(* Logix 5000 project; controller MV vendor 1 type 14 code 217 rev 31.11; software revision 31.00; part 9 of 53 *)
(* tags used below, declared in another part *)
   MC_CH1_DRAIN : PlantItem;   // CH1_DRAIN
   MC_CH1_LF1 : PlantItem;   // CH1_LF1
   MC_CH1_PR1 : PlantItem;   // CH1_PR1
   MC_CH1_RR : PlantItem;   // CH1_RR
   MC_N100 : INT[255];   // C1_PLC Channel 1 PLC data
   MC_N102 : INT[255];   // CH1 PROG Channel 1 CIP progra m
   MC_N104 : INT[255];   // CH1 REPORT Channel 1 CIP report file
   MC_N112 : INT[255];   // FVR DATA Data read from FV ro uting PLC
   MC_N113 : INT[255];   // MVR DATA Data read from MV ro uting PLC
   MC_N114 : INT[255];   // YP DATA
   MC_N120 : INT[255];   // C2 PLC Channel 2 PLC data
   MC_N80 : INT[255];   // SRV1_PLC Detergent tank 1 ser vice PLC data
   MC_N90 : INT[255];   // SV2_PLC Detergent tank 2 ser vice PLC data
   MC_T105 : TIMER[255];   // CH1 TIMERS Channel 1 timers
   MC_T4 : TIMER[255];   // TIMER
(* MC_Common, continued *)

ROUTINE MC_CH1_POSTRN_113   (* ladder *)
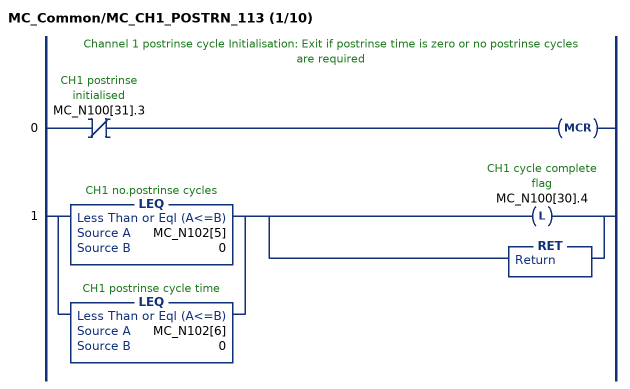
   // Channel 1 postrinse cycle Initialisation: Exit if postrinse time is zero or no postrinse cycles are required
   0: XIO(MC_N100[31].3)MCR();
   1: [LEQ(MC_N102[5],0) ,LEQ(MC_N102[6],0) ][OTL(MC_N100[30].4) ,RET() ];
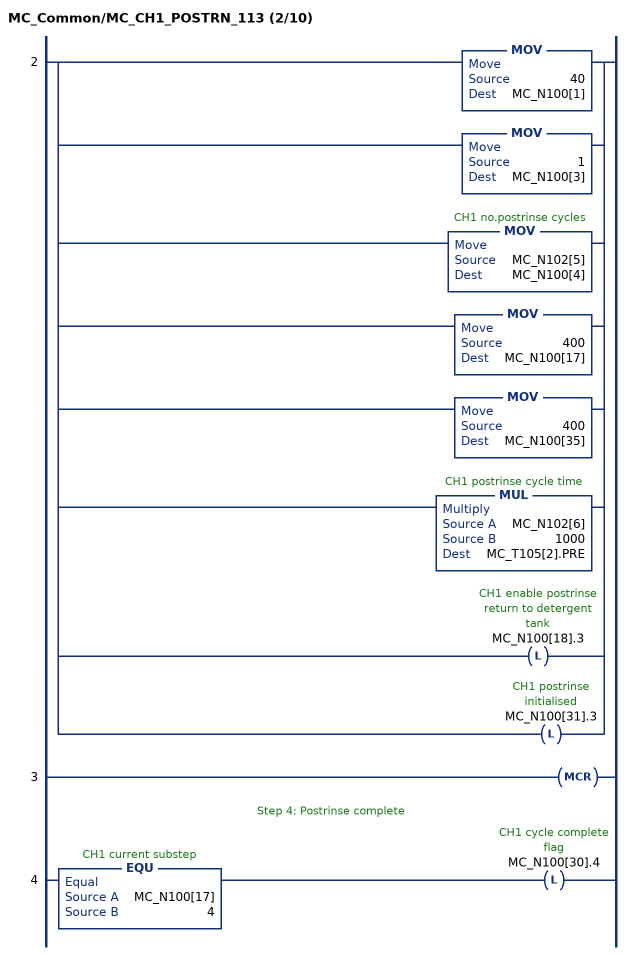
   2: [MOV(40,MC_N100[1]) ,MOV(1,MC_N100[3]) ,MOV(MC_N102[5],MC_N100[4]) ,MOV(400,MC_N100[17]) ,MOV(400,MC_N100[35]) ,MUL(MC_N102[6],1000,MC_T105[2].PRE) ,OTL(MC_N100[18].3) ,OTL(MC_N100[31].3) ];
   3: MCR();
   // Step 4: Postrinse complete
   4: EQU(MC_N100[17],4)OTL(MC_N100[30].4);
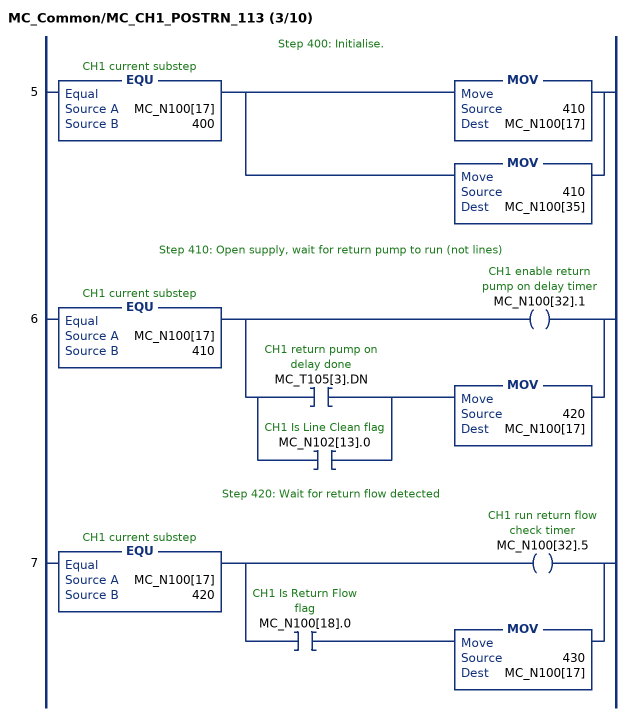
   // Step 400: Initialise.
   5: EQU(MC_N100[17],400)[MOV(410,MC_N100[17]) ,MOV(410,MC_N100[35]) ];
   // Step 410: Open supply, wait for return pump to run (not lines)
   6: EQU(MC_N100[17],410)[OTE(MC_N100[32].1) ,[XIC(MC_T105[3].DN) ,XIC(MC_N102[13].0) ] MOV(420,MC_N100[17]) ];
   // Step 420: Wait for return flow detected
   7: EQU(MC_N100[17],420)[OTE(MC_N100[32].5) ,XIC(MC_N100[18].0) MOV(430,MC_N100[17]) ];
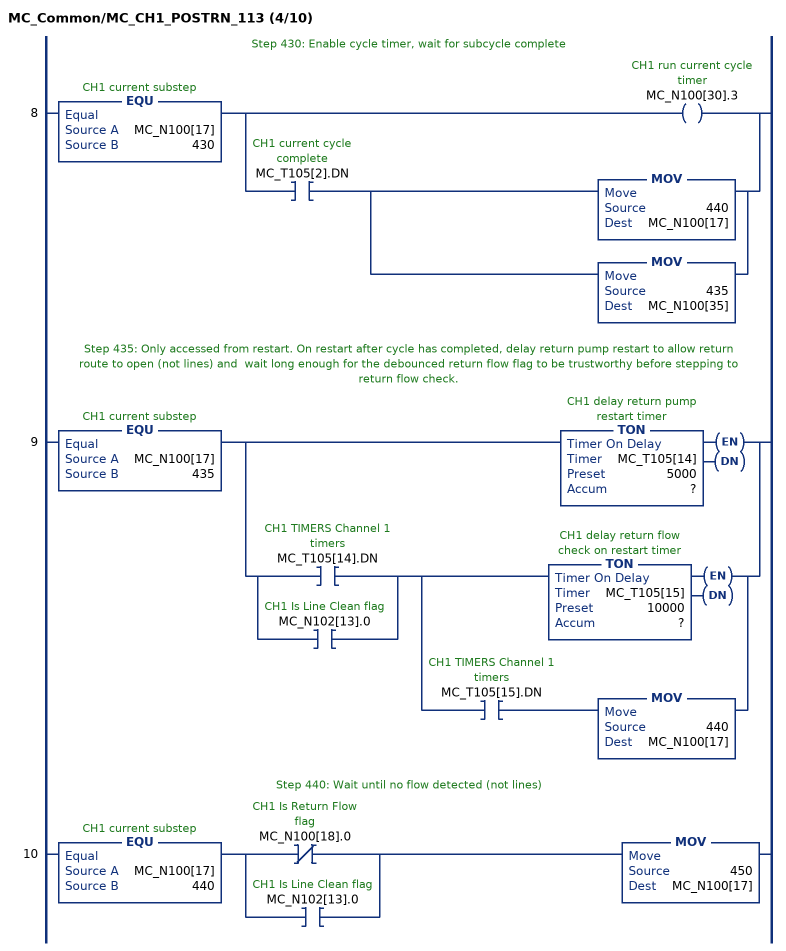
   // Step 430: Enable cycle timer, wait for subcycle complete
   8: EQU(MC_N100[17],430)[OTE(MC_N100[30].3) ,XIC(MC_T105[2].DN) [MOV(440,MC_N100[17]) ,MOV(435,MC_N100[35]) ] ];
   // Step 435: Only accessed from restart. On restart after cycle has completed, delay return pump restart to allow return route to open (not lines) and  wait long enough for the debounced return flow flag to be trustworthy before stepping to return flow check.
   9: EQU(MC_N100[17],435)[TON(MC_T105[14],?,?) ,[XIC(MC_T105[14].DN) ,XIC(MC_N102[13].0) ] [TON(MC_T105[15],?,?) ,XIC(MC_T105[15].DN) MOV(440,MC_N100[17]) ] ];
   // Step 440: Wait until no flow detected (not lines)
   10: EQU(MC_N100[17],440)[XIO(MC_N100[18].0) ,XIC(MC_N102[13].0) ]MOV(450,MC_N100[17]);
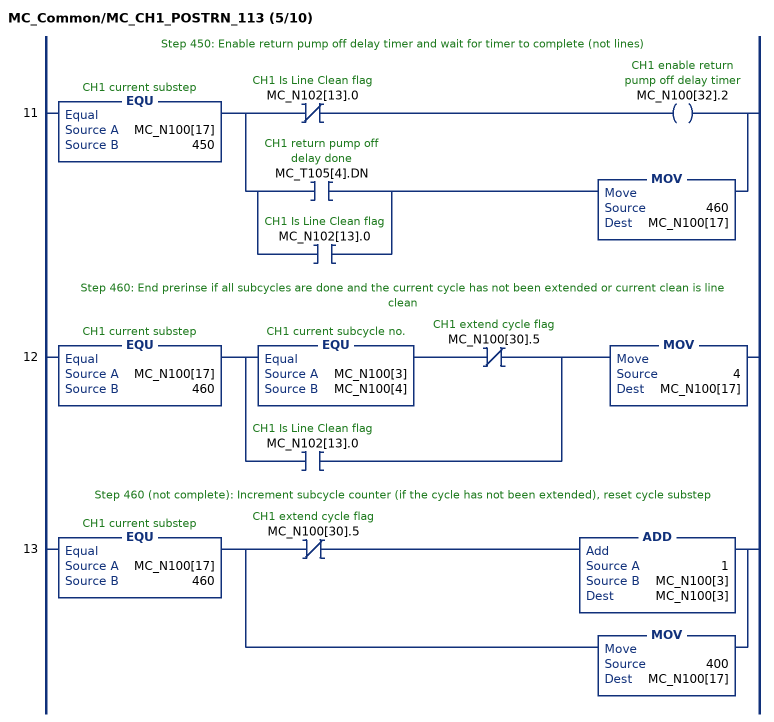
   // Step 450: Enable return pump off delay timer and wait for timer to complete (not lines)
   11: EQU(MC_N100[17],450)[XIO(MC_N102[13].0) OTE(MC_N100[32].2) ,[XIC(MC_T105[4].DN) ,XIC(MC_N102[13].0) ] MOV(460,MC_N100[17]) ];
   // Step 460: End prerinse if all subcycles are done and the current cycle has not been extended or current clean is line clean
   12: EQU(MC_N100[17],460)[EQU(MC_N100[3],MC_N100[4]) XIO(MC_N100[30].5) ,XIC(MC_N102[13].0) ]MOV(4,MC_N100[17]);
   // Step 460 (not complete): Increment subcycle counter (if the cycle has not been extended), reset cycle substep
   13: EQU(MC_N100[17],460)[XIO(MC_N100[30].5) ADD(1,MC_N100[3],MC_N100[3]) ,MOV(400,MC_N100[17]) ];
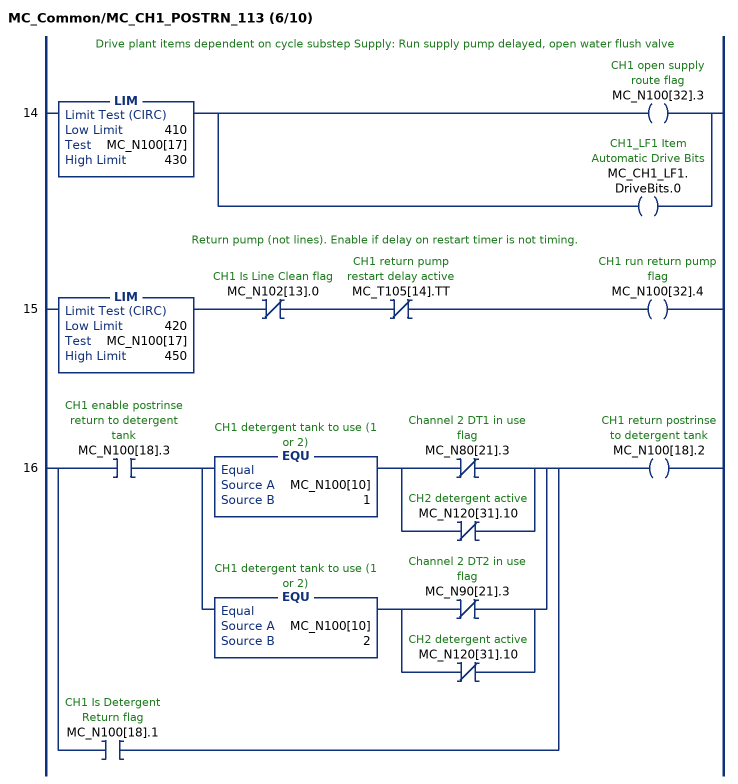
   // Drive plant items dependent on cycle substep Supply: Run supply pump delayed, open water flush valve
   14: LIM(410,MC_N100[17],430)[OTE(MC_N100[32].3) ,OTE(MC_CH1_LF1.DriveBits.0) ];
   // Return pump (not lines). Enable if delay on restart timer is not timing.
   15: LIM(420,MC_N100[17],450)XIO(MC_N102[13].0)XIO(MC_T105[14].TT)OTE(MC_N100[32].4);
   16: [XIC(MC_N100[18].3) [EQU(MC_N100[10],1) [XIO(MC_N80[21].3) ,XIO(MC_N120[31].10) ] ,EQU(MC_N100[10],2) [XIO(MC_N90[21].3) ,XIO(MC_N120[31].10) ] ] ,XIC(MC_N100[18].1) ]OTE(MC_N100[18].2);
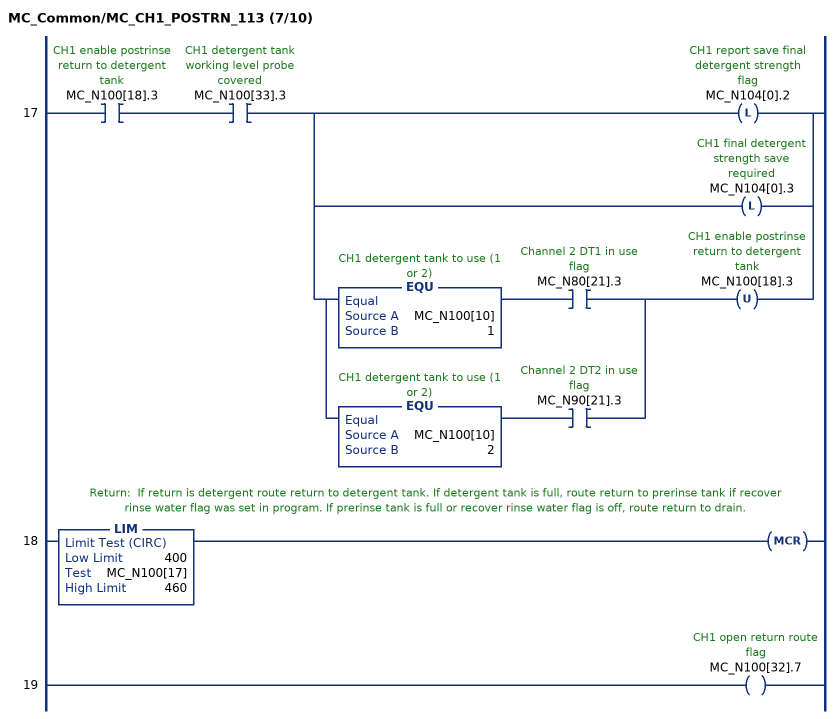
   17: XIC(MC_N100[18].3)XIC(MC_N100[33].3)[OTL(MC_N104[0].2) ,OTL(MC_N104[0].3) ,[EQU(MC_N100[10],1) XIC(MC_N80[21].3) ,EQU(MC_N100[10],2) XIC(MC_N90[21].3) ] OTU(MC_N100[18].3) ];
   // Return:  If return is detergent route return to detergent tank. If detergent tank is full, route return to prerinse tank if recover rinse water flag was set in program. If prerinse tank is full or recover rinse water flag is off, route return to drain.
   18: LIM(400,MC_N100[17],460)MCR();
   19: OTE(MC_N100[32].7);
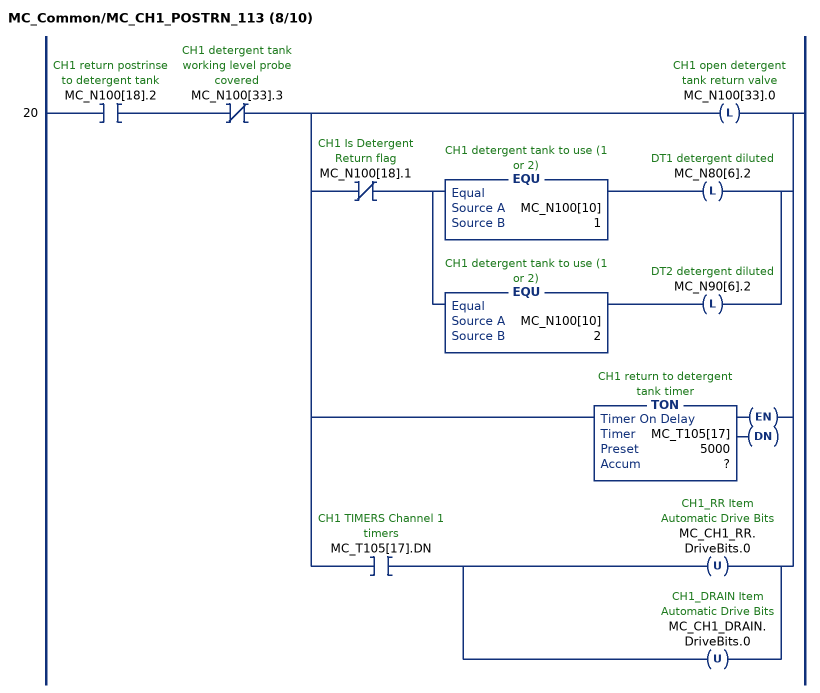
   20: XIC(MC_N100[18].2)XIO(MC_N100[33].3)[OTL(MC_N100[33].0) ,XIO(MC_N100[18].1) [EQU(MC_N100[10],1) OTL(MC_N80[6].2) ,EQU(MC_N100[10],2) OTL(MC_N90[6].2) ] ,TON(MC_T105[17],?,?) ,XIC(MC_T105[17].DN) [OTU(MC_CH1_RR.DriveBits.0) ,OTU(MC_CH1_DRAIN.DriveBits.0) ] ];
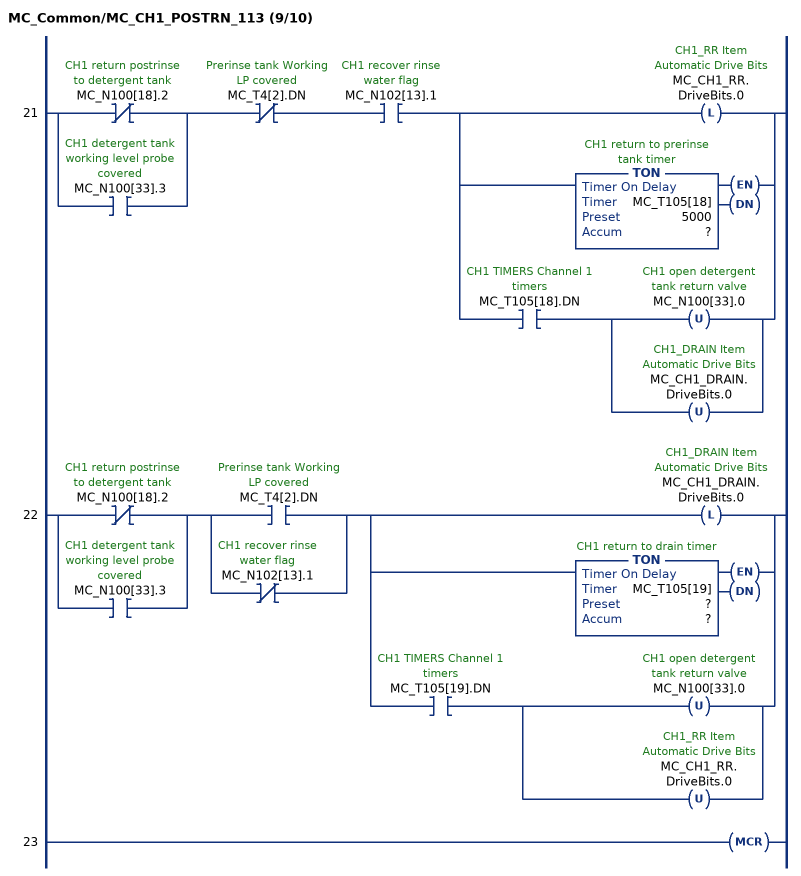
   21: [XIO(MC_N100[18].2) ,XIC(MC_N100[33].3) ]XIO(MC_T4[2].DN)XIC(MC_N102[13].1)[OTL(MC_CH1_RR.DriveBits.0) ,TON(MC_T105[18],?,?) ,XIC(MC_T105[18].DN) [OTU(MC_N100[33].0) ,OTU(MC_CH1_DRAIN.DriveBits.0) ] ];
   22: [XIO(MC_N100[18].2) ,XIC(MC_N100[33].3) ][XIC(MC_T4[2].DN) ,XIO(MC_N102[13].1) ][OTL(MC_CH1_DRAIN.DriveBits.0) ,TON(MC_T105[19],?,?) ,XIC(MC_T105[19].DN) [OTU(MC_N100[33].0) ,OTU(MC_CH1_RR.DriveBits.0) ] ];
   23: MCR();
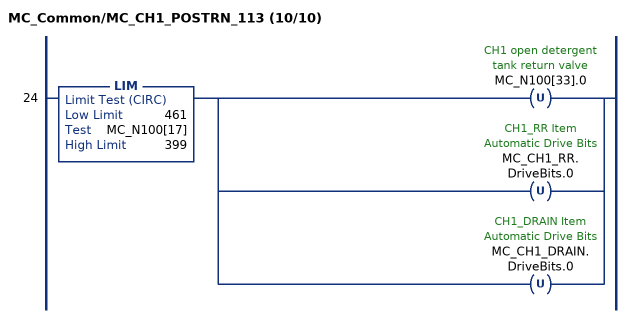
   24: LIM(461,MC_N100[17],399)[OTU(MC_N100[33].0) ,OTU(MC_CH1_RR.DriveBits.0) ,OTU(MC_CH1_DRAIN.DriveBits.0) ];
END_ROUTINE

ROUTINE MC_CH1_PRERN_111   (* ladder *)
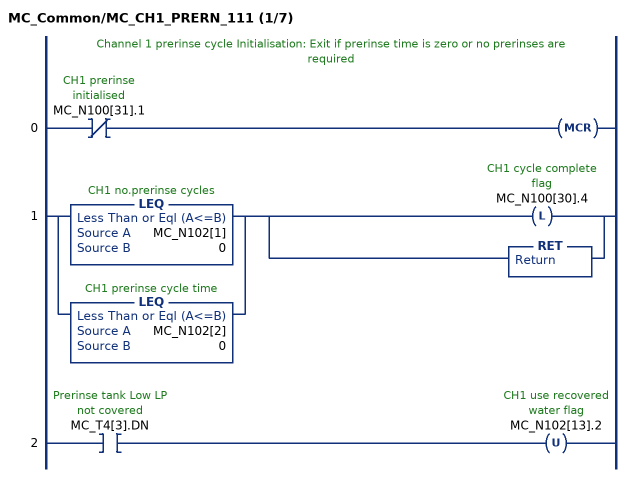
   // Channel 1 prerinse cycle Initialisation: Exit if prerinse time is zero or no prerinses are required
   0: XIO(MC_N100[31].1)MCR();
   1: [LEQ(MC_N102[1],0) ,LEQ(MC_N102[2],0) ][OTL(MC_N100[30].4) ,RET() ];
   2: XIC(MC_T4[3].DN)OTU(MC_N102[13].2);
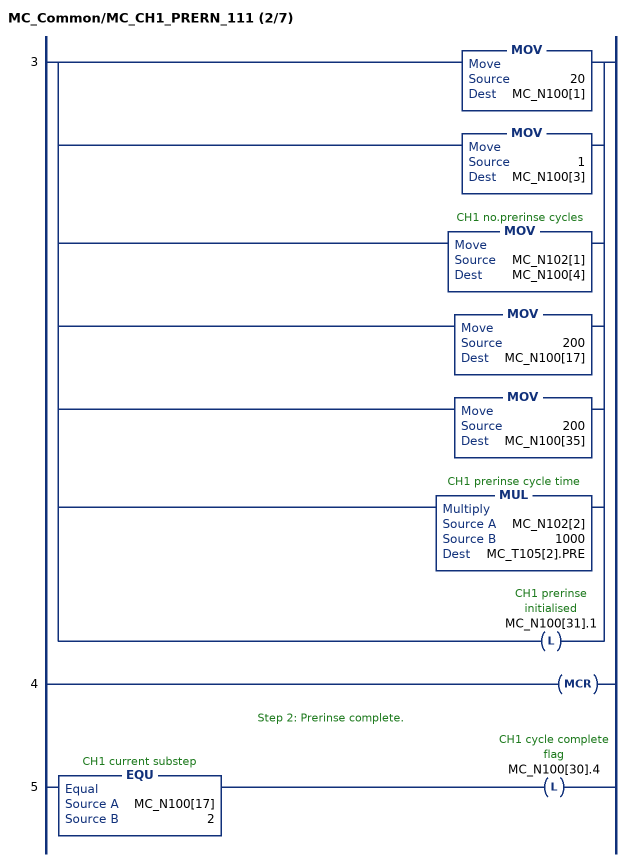
   3: [MOV(20,MC_N100[1]) ,MOV(1,MC_N100[3]) ,MOV(MC_N102[1],MC_N100[4]) ,MOV(200,MC_N100[17]) ,MOV(200,MC_N100[35]) ,MUL(MC_N102[2],1000,MC_T105[2].PRE) ,OTL(MC_N100[31].1) ];
   4: MCR();
   // Step 2: Prerinse complete.
   5: EQU(MC_N100[17],2)OTL(MC_N100[30].4);
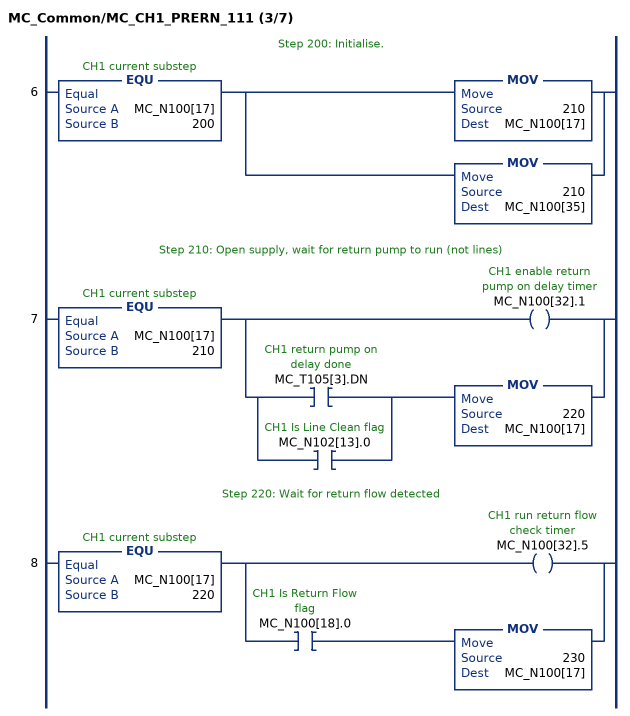
   // Step 200: Initialise.
   6: EQU(MC_N100[17],200)[MOV(210,MC_N100[17]) ,MOV(210,MC_N100[35]) ];
   // Step 210: Open supply, wait for return pump to run (not lines)
   7: EQU(MC_N100[17],210)[OTE(MC_N100[32].1) ,[XIC(MC_T105[3].DN) ,XIC(MC_N102[13].0) ] MOV(220,MC_N100[17]) ];
   // Step 220: Wait for return flow detected
   8: EQU(MC_N100[17],220)[OTE(MC_N100[32].5) ,XIC(MC_N100[18].0) MOV(230,MC_N100[17]) ];
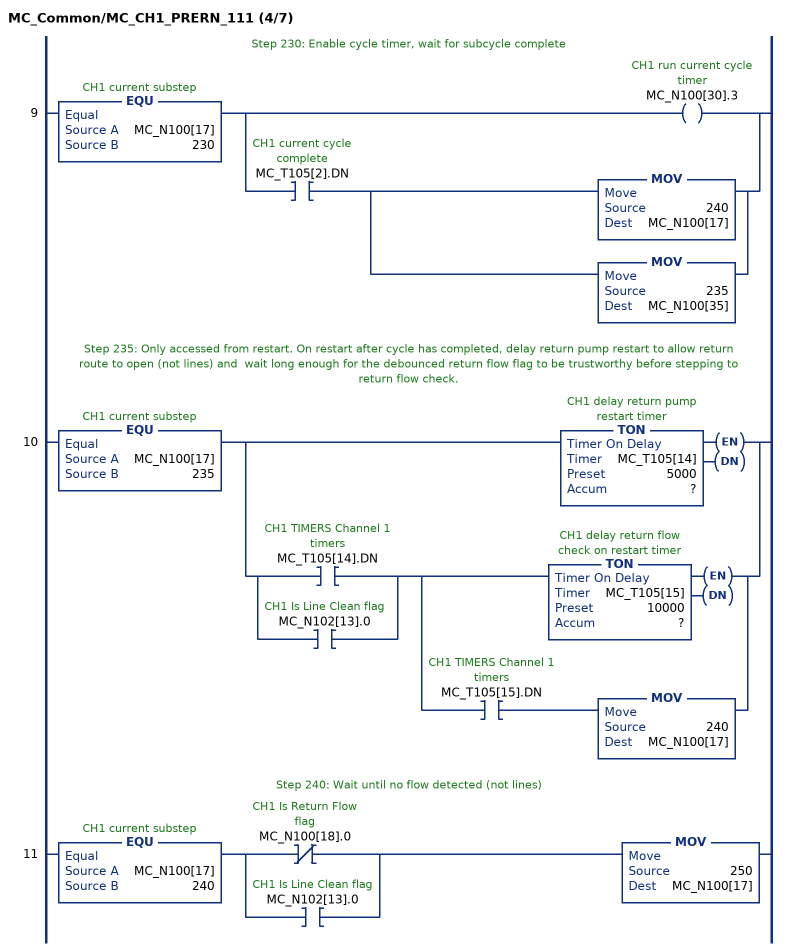
   // Step 230: Enable cycle timer, wait for subcycle complete
   9: EQU(MC_N100[17],230)[OTE(MC_N100[30].3) ,XIC(MC_T105[2].DN) [MOV(240,MC_N100[17]) ,MOV(235,MC_N100[35]) ] ];
   // Step 235: Only accessed from restart. On restart after cycle has completed, delay return pump restart to allow return route to open (not lines) and  wait long enough for the debounced return flow flag to be trustworthy before stepping to return flow check.
   10: EQU(MC_N100[17],235)[TON(MC_T105[14],?,?) ,[XIC(MC_T105[14].DN) ,XIC(MC_N102[13].0) ] [TON(MC_T105[15],?,?) ,XIC(MC_T105[15].DN) MOV(240,MC_N100[17]) ] ];
   // Step 240: Wait until no flow detected (not lines)
   11: EQU(MC_N100[17],240)[XIO(MC_N100[18].0) ,XIC(MC_N102[13].0) ]MOV(250,MC_N100[17]);
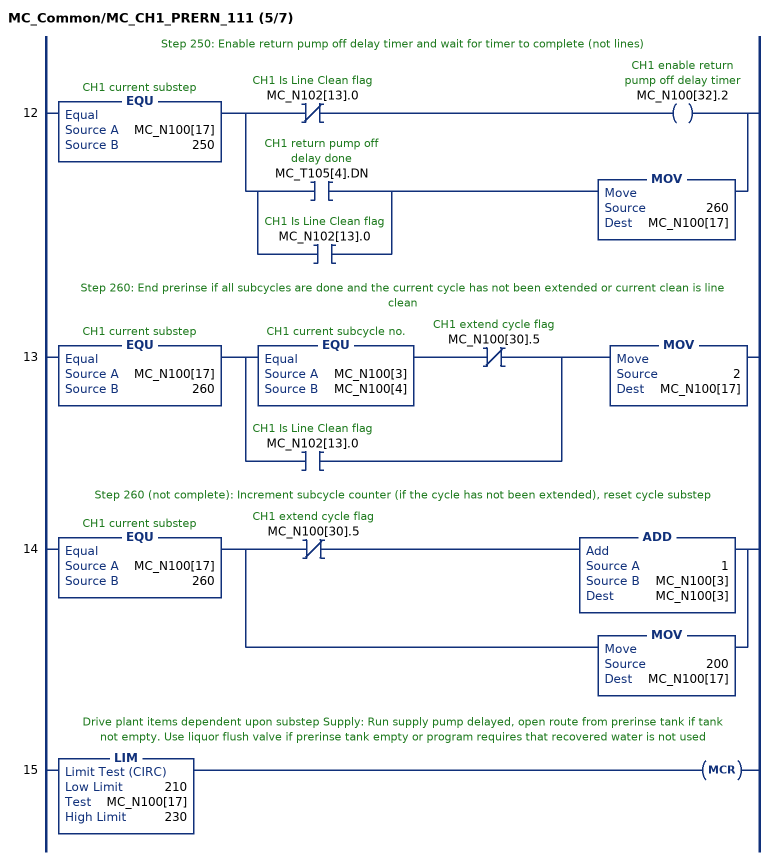
   // Step 250: Enable return pump off delay timer and wait for timer to complete (not lines)
   12: EQU(MC_N100[17],250)[XIO(MC_N102[13].0) OTE(MC_N100[32].2) ,[XIC(MC_T105[4].DN) ,XIC(MC_N102[13].0) ] MOV(260,MC_N100[17]) ];
   // Step 260: End prerinse if all subcycles are done and the current cycle has not been extended or current clean is line clean
   13: EQU(MC_N100[17],260)[EQU(MC_N100[3],MC_N100[4]) XIO(MC_N100[30].5) ,XIC(MC_N102[13].0) ]MOV(2,MC_N100[17]);
   // Step 260 (not complete): Increment subcycle counter (if the cycle has not been extended), reset cycle substep
   14: EQU(MC_N100[17],260)[XIO(MC_N100[30].5) ADD(1,MC_N100[3],MC_N100[3]) ,MOV(200,MC_N100[17]) ];
   // Drive plant items dependent upon substep Supply: Run supply pump delayed, open route from prerinse tank if tank not empty. Use liquor flush valve if prerinse tank empty or program requires that recovered water is not used
   15: LIM(210,MC_N100[17],230)MCR();
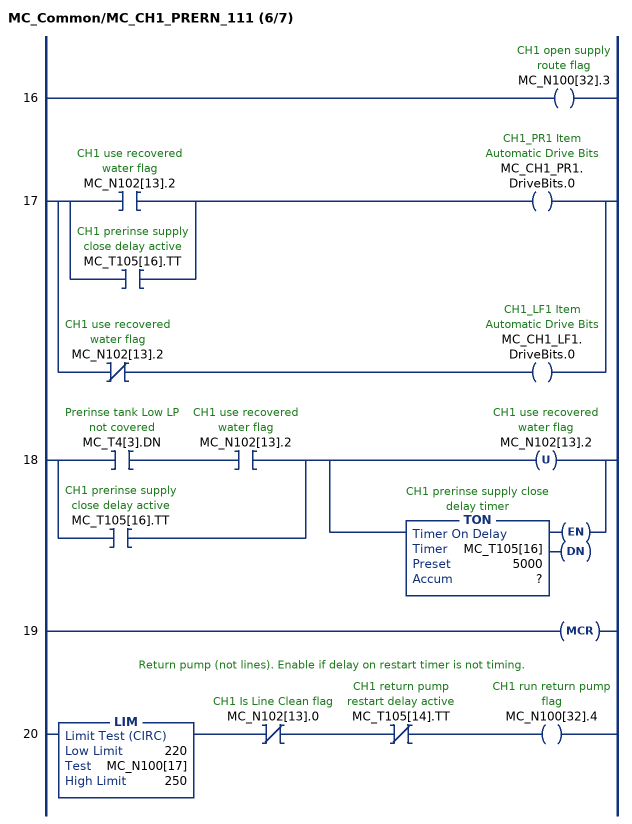
   16: OTE(MC_N100[32].3);
   17: [[XIC(MC_N102[13].2) ,XIC(MC_T105[16].TT) ] OTE(MC_CH1_PR1.DriveBits.0) ,XIO(MC_N102[13].2) OTE(MC_CH1_LF1.DriveBits.0) ];
   18: [XIC(MC_T4[3].DN) XIC(MC_N102[13].2) ,XIC(MC_T105[16].TT) ][OTU(MC_N102[13].2) ,TON(MC_T105[16],?,?) ];
   19: MCR();
   // Return pump (not lines). Enable if delay on restart timer is not timing.
   20: LIM(220,MC_N100[17],250)XIO(MC_N102[13].0)XIO(MC_T105[14].TT)OTE(MC_N100[32].4);
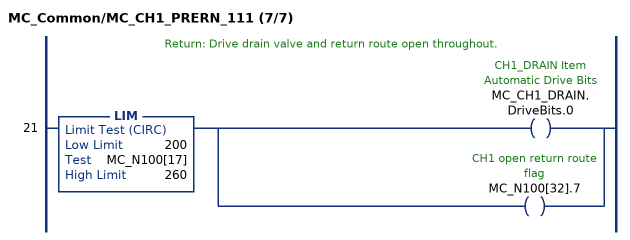
   // Return: Drive drain valve and return route open throughout.
   21: LIM(200,MC_N100[17],260)[OTE(MC_CH1_DRAIN.DriveBits.0) ,OTE(MC_N100[32].7) ];
END_ROUTINE

ROUTINE MC_CH1_REPORT_104   (* ladder *)
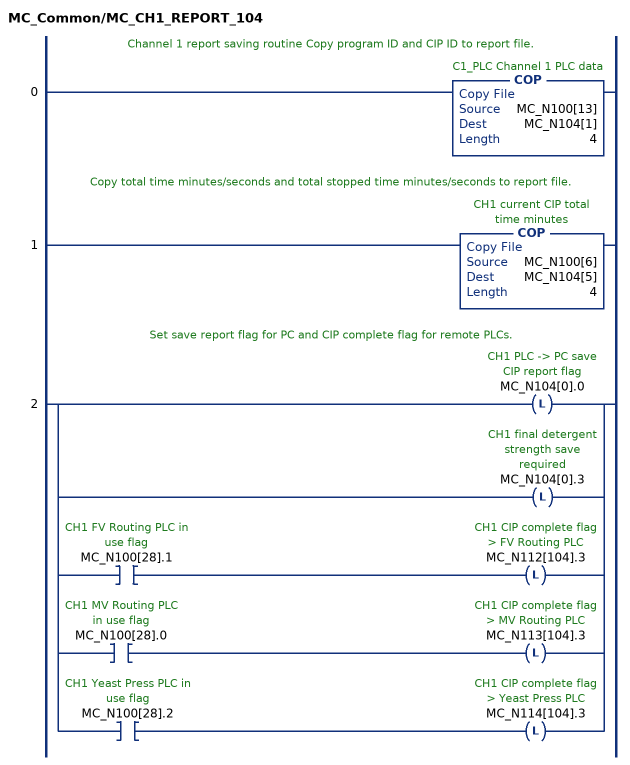
   // Channel 1 report saving routine Copy program ID and CIP ID to report file.
   0: COP(MC_N100[13],MC_N104[1],4);
   // Copy total time minutes/seconds and total stopped time minutes/seconds to report file.
   1: COP(MC_N100[6],MC_N104[5],4);
   // Set save report flag for PC and CIP complete flag for remote PLCs.
   2: [OTL(MC_N104[0].0) ,OTL(MC_N104[0].3) ,XIC(MC_N100[28].1) OTL(MC_N112[104].3) ,XIC(MC_N100[28].0) OTL(MC_N113[104].3) ,XIC(MC_N100[28].2) OTL(MC_N114[104].3) ];
END_ROUTINE
